(* Logix 5000 project; controller FV vendor 1 type 14 code 217 rev 31.11; software revision 31.00; part 27 of 63 *)
(* tags used below, declared in another part *)
   Alarm_Reset : BOOL;
   Default_Check_Time : DINT;
   Dummy : BOOL;
   FR_B230 : INT[255];   // FLOW_BITS Flow Meter Bits
   FR_B240 : INT[255];   // DEBOUNCE Debounce Flags
   FR_B246 : INT[255];   // V_REVERSE Flags for reversing contol action
   FR_B247 : INT[255];   // CHECKWORD Simulation Flags for Checkwords
   FR_B248 : INT[255];   // FORCE ON Force On Flags
   FR_B249 : INT[255];   // FORCE_OFF NOT Force Off Flags
   FR_B3 : INT[255];   // BINARY
   FR_bit_data_file_address : DINT;
   FR_bit_file_bit_offset : DINT;
   FR_bit_file_word_offset : DINT;
   FR_bit_offset : DINT;
   FR_bit_value_to_set : DINT;
   FR_data_file_address : DINT;
   FR_FRV1_AV01 : PlantItem;   // FRV1_AV01
   FR_FRV1_AV01_ALARM : ALARM_DIGITAL;
   FR_FRV1_AV01_C : ALIAS FOR RIO_Rack_2:4:I.Data.15;
   FR_FRV1_AV01_DR : ALIAS FOR RIO_Rack_2:5:O.Data.7;
   FR_FRV1_AV01_O : ALIAS FOR RIO_Rack_2:4:I.Data.11;
   FR_FV26_AV01 : PlantItem;   // FV26_AV01
   FR_FV26_AV01_ALARM : ALARM_DIGITAL;
   FR_FV26_AV01_C : ALIAS FOR RIO_Rack_2:4:I.Data.20;
   FR_FV26_AV01_O : ALIAS FOR RIO_Rack_2:4:I.Data.16;
   FR_FV26_AV01_RDR : ALIAS FOR RIO_Rack_2:5:O.Data.8;
   FR_FV26_AV04 : PlantItem;   // FV26_AV04
   FR_FV26_AV04_ALARM : ALARM_DIGITAL;
   FR_FV26_AV04_C : ALIAS FOR RIO_Rack_2:4:I.Data.21;
   FR_FV26_AV04_DR : ALIAS FOR RIO_Rack_2:5:O.Data.9;
   FR_FV26_AV04_O : ALIAS FOR RIO_Rack_2:4:I.Data.17;
   FR_FV26_AV05 : PlantItem;   // FV26_AV05
   FR_FV26_AV05_ALARM : ALARM_DIGITAL;
   FR_FV26_AV05_C : ALIAS FOR RIO_Rack_2:4:I.Data.22;
   FR_FV26_AV05_DR : ALIAS FOR RIO_Rack_2:5:O.Data.10;
   FR_FV26_AV05_O : ALIAS FOR RIO_Rack_2:4:I.Data.18;
   FR_FV26_AV06 : PlantItem;   // FV26_AV06
   FR_FV26_AV06_ALARM : ALARM_DIGITAL;
   FR_FV26_AV06_C : ALIAS FOR RIO_Rack_2:4:I.Data.23;
   FR_FV26_AV06_DR : ALIAS FOR RIO_Rack_2:5:O.Data.11;
   FR_FV26_AV06_O : ALIAS FOR RIO_Rack_2:4:I.Data.19;
   FR_FV26_AV07 : PlantItem;   // FV26_AV07
   FR_FV26_AV07_ALARM : ALARM_DIGITAL;
   FR_FV26_AV07_C : ALIAS FOR RIO_Rack_2:4:I.Data.28;
   FR_FV26_AV07_DR : ALIAS FOR RIO_Rack_2:5:O.Data.12;
   FR_FV26_AV07_O : ALIAS FOR RIO_Rack_2:4:I.Data.24;
   FR_FV27_AV01 : PlantItem;   // FV27_AV01
   FR_FV27_AV01_ALARM : ALARM_DIGITAL;
   FR_FV27_AV01_C : ALIAS FOR RIO_Rack_2:4:I.Data.29;
   FR_FV27_AV01_O : ALIAS FOR RIO_Rack_2:4:I.Data.25;
   FR_FV27_AV01_RDR : ALIAS FOR RIO_Rack_2:5:O.Data.13;
   FR_FV27_AV04 : PlantItem;   // FV27_AV04
   FR_FV27_AV04_ALARM : ALARM_DIGITAL;
   FR_FV27_AV04_C : ALIAS FOR RIO_Rack_2:4:I.Data.30;
   FR_FV27_AV04_DR : ALIAS FOR RIO_Rack_2:5:O.Data.14;
   FR_FV27_AV04_O : ALIAS FOR RIO_Rack_2:4:I.Data.26;
   FR_FV27_AV05 : PlantItem;   // FV27_AV05
   FR_FV27_AV05_ALARM : ALARM_DIGITAL;
   FR_FV27_AV05_C : ALIAS FOR RIO_Rack_2:4:I.Data.31;
   FR_FV27_AV05_DR : ALIAS FOR RIO_Rack_2:5:O.Data.15;
   FR_FV27_AV05_O : ALIAS FOR RIO_Rack_2:4:I.Data.27;
   FR_FV27_AV06 : PlantItem;   // FV27_AV06
   FR_FV27_AV06_ALARM : ALARM_DIGITAL;
   FR_FV27_AV06_C : ALIAS FOR RIO_Rack_2:6:I.Data.4;
   FR_FV27_AV06_DR : ALIAS FOR RIO_Rack_2:5:O.Data.16;
   FR_FV27_AV06_O : ALIAS FOR RIO_Rack_2:6:I.Data.0;
   FR_FV27_AV07 : PlantItem;   // FV27_AV07
   FR_FV27_AV07_ALARM : ALARM_DIGITAL;
   FR_FV27_AV07_C : ALIAS FOR RIO_Rack_2:6:I.Data.5;
   FR_FV27_AV07_DR : ALIAS FOR RIO_Rack_2:5:O.Data.17;
   FR_FV27_AV07_O : ALIAS FOR RIO_Rack_2:6:I.Data.1;
   FR_N10 : INT[265];   // FV_AGING Comms to FV Aging PL C
   FR_N100 : INT[265];   // FV FILLING
   FR_N110 : INT[265];   // GREEN BEER Green Beer Main
   FR_N120 : INT[265];   // YEAST CROP Yeast Cropping Main
   FR_N13 : INT[265];   // MV_ROUTE Comms to MV Routing PLC
   FR_N130 : INT[265];   // FILTRATE Filtrate Return
   FR_N14 : INT[265];   // MVFV CIP Comms to MVFV CIP Un it PLC
   FR_N140 : INT[265];   // CIP
   FR_N142 : INT[265];   // CIP
   FR_N143 : INT[265];   // CIP
   FR_N150 : INT[265];   // Original N File From SLC, No Description Available
   FR_N160 : INT[265];   // VESSEL Vessel Working Direc tory
   FR_N170 : INT[265];   // Original N File From SLC, No Description Available
   FR_N180 : INT[265];   // Original N File From SLC, No Description Available
   FR_N198 : INT[265];   // Original N File From SLC, No Description Available
   FR_N20 : INT[265];   // GENERAL General Purpose Setp oints
   FR_N200 : INT[265];   // ANALOG_IN Analog Inputs
   FR_N201 : INT[265];   // Original N File From SLC, No Description Available
   FR_N207 : INT[265];   // Original N File From SLC, No Description Available
   FR_N21 : INT[265];   // CHASE_V FV Filling Beer Chas e Volumes
   FR_N210 : INT[265];   // ANALOG_OUT Analog Outputs
   FR_N220 : INT[265];   // CHECKLIST Checklist Loop Contr ollers
   FR_N225 : INT[265];   // Original N File From SLC, No Description Available
   FR_N226 : INT[265];   // Original N File From SLC, No Description Available
   FR_N245 : INT[265];   // CHECKWORD Checkword Loop Contr ol
   FR_N252 : INT[265];   // OUTPUT_PTR Checkword Pointers t o output flags in B2 50
   FR_N253 : INT[265];   // EN_POINT Pointers to energise d input flags in B25 1
   FR_N254 : INT[265];   // DEN_POINT Pointers to deenergi sed input flags in B 251
   FR_N255 : INT[265];   // CHECKWORDS
   FR_N26 : INT[265];   // FV26
   FR_N27 : INT[265];   // FV27
   FR_N28 : INT[265];   // FV28
   FR_N29 : INT[265];   // FV29
   FR_N30 : INT[265];   // FV30
   FR_N31 : INT[265];   // FV31
   FR_N36 : INT[265];   // Original N File From SLC, No Description Available
   FR_N37 : INT[265];   // Original N File From SLC, No Description Available
   FR_N46 : INT[265];   // Original N File From SLC, No Description Available
   FR_N47 : INT[265];   // Original N File From SLC, No Description Available
   FR_N7 : INT[265];   // INTEGER
   FR_N99 : INT[265];   // COMMENT Comment Lines
   FR_value_to_set : DINT;
   FR_VB1_AV01 : PlantItem;   // VB1_AV01
   FR_VB1_AV01_ALARM : ALARM_DIGITAL;
   FR_VB1_AV01_C : ALIAS FOR RIO_Rack_2:6:I.Data.6;
   FR_VB1_AV01_DR : ALIAS FOR RIO_Rack_2:5:O.Data.18;
   FR_VB1_AV01_O : ALIAS FOR RIO_Rack_2:6:I.Data.2;
   FR_VB1_AV02 : PlantItem;   // VB1_AV02
   FR_VB1_AV02_ALARM : ALARM_DIGITAL;
   FR_VB1_AV02_C : ALIAS FOR RIO_Rack_2:6:I.Data.7;
   FR_VB1_AV02_DR : ALIAS FOR RIO_Rack_2:5:O.Data.19;
   FR_VB1_AV02_O : ALIAS FOR RIO_Rack_2:6:I.Data.3;
   FR_VB1_AV03 : PlantItem;   // VB1_AV03
   FR_VB1_AV03_ALARM : ALARM_DIGITAL;
   FR_VB1_AV03_C : ALIAS FOR RIO_Rack_2:6:I.Data.12;
   FR_VB1_AV03_DR : ALIAS FOR RIO_Rack_2:5:O.Data.20;
   FR_VB1_AV03_O : ALIAS FOR RIO_Rack_2:6:I.Data.8;
   FR_word_offset : DINT;
   Item_Faults_Are_Latched : BOOL;
   Item_Simulation_Flag : BOOL;
   One_Second_One_Scan : ALIAS FOR One_Second_1_scan;
(* FR_Common, continued *)

ROUTINE FR_Set_NFile_Value   (* ladder *)
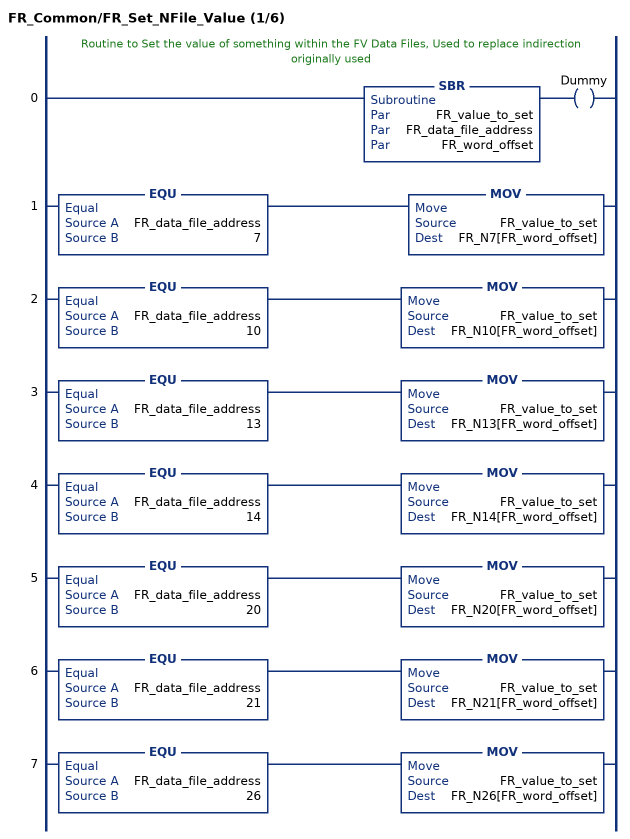
   // Routine to Set the value of something within the FV Data Files, Used to replace indirection originally used
   0: SBR(FR_value_to_set,FR_data_file_address,FR_word_offset)OTE(Dummy);
   1: EQU(FR_data_file_address,7)MOV(FR_value_to_set,FR_N7[FR_word_offset]);
   2: EQU(FR_data_file_address,10)MOV(FR_value_to_set,FR_N10[FR_word_offset]);
   3: EQU(FR_data_file_address,13)MOV(FR_value_to_set,FR_N13[FR_word_offset]);
   4: EQU(FR_data_file_address,14)MOV(FR_value_to_set,FR_N14[FR_word_offset]);
   5: EQU(FR_data_file_address,20)MOV(FR_value_to_set,FR_N20[FR_word_offset]);
   6: EQU(FR_data_file_address,21)MOV(FR_value_to_set,FR_N21[FR_word_offset]);
   7: EQU(FR_data_file_address,26)MOV(FR_value_to_set,FR_N26[FR_word_offset]);
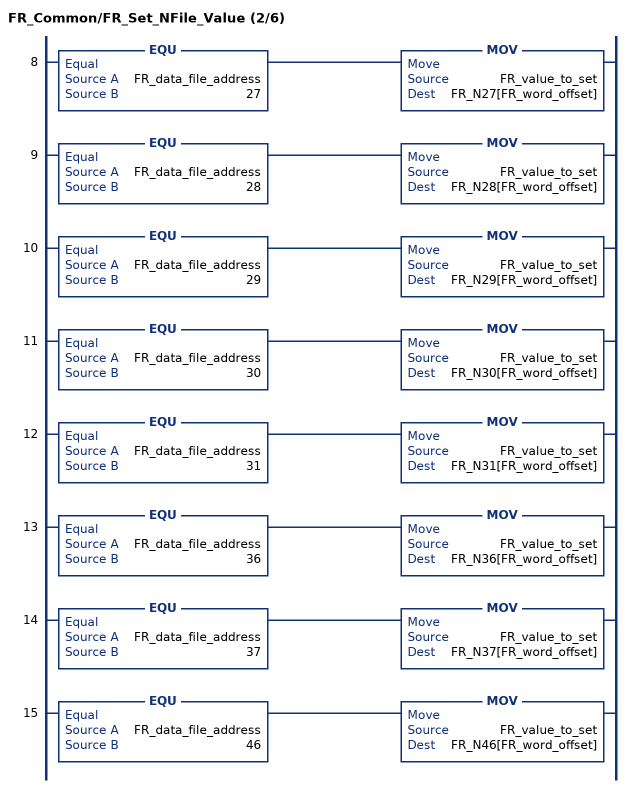
   8: EQU(FR_data_file_address,27)MOV(FR_value_to_set,FR_N27[FR_word_offset]);
   9: EQU(FR_data_file_address,28)MOV(FR_value_to_set,FR_N28[FR_word_offset]);
   10: EQU(FR_data_file_address,29)MOV(FR_value_to_set,FR_N29[FR_word_offset]);
   11: EQU(FR_data_file_address,30)MOV(FR_value_to_set,FR_N30[FR_word_offset]);
   12: EQU(FR_data_file_address,31)MOV(FR_value_to_set,FR_N31[FR_word_offset]);
   13: EQU(FR_data_file_address,36)MOV(FR_value_to_set,FR_N36[FR_word_offset]);
   14: EQU(FR_data_file_address,37)MOV(FR_value_to_set,FR_N37[FR_word_offset]);
   15: EQU(FR_data_file_address,46)MOV(FR_value_to_set,FR_N46[FR_word_offset]);
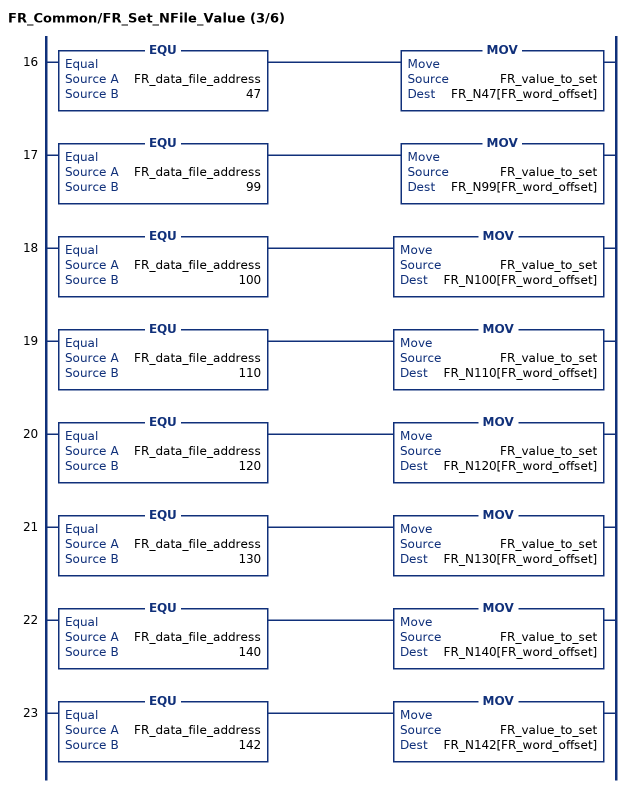
   16: EQU(FR_data_file_address,47)MOV(FR_value_to_set,FR_N47[FR_word_offset]);
   17: EQU(FR_data_file_address,99)MOV(FR_value_to_set,FR_N99[FR_word_offset]);
   18: EQU(FR_data_file_address,100)MOV(FR_value_to_set,FR_N100[FR_word_offset]);
   19: EQU(FR_data_file_address,110)MOV(FR_value_to_set,FR_N110[FR_word_offset]);
   20: EQU(FR_data_file_address,120)MOV(FR_value_to_set,FR_N120[FR_word_offset]);
   21: EQU(FR_data_file_address,130)MOV(FR_value_to_set,FR_N130[FR_word_offset]);
   22: EQU(FR_data_file_address,140)MOV(FR_value_to_set,FR_N140[FR_word_offset]);
   23: EQU(FR_data_file_address,142)MOV(FR_value_to_set,FR_N142[FR_word_offset]);
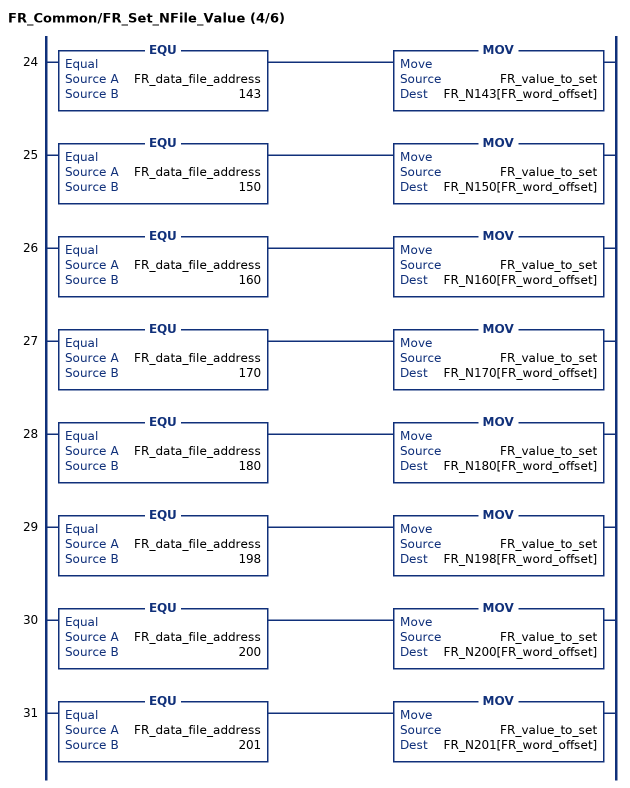
   24: EQU(FR_data_file_address,143)MOV(FR_value_to_set,FR_N143[FR_word_offset]);
   25: EQU(FR_data_file_address,150)MOV(FR_value_to_set,FR_N150[FR_word_offset]);
   26: EQU(FR_data_file_address,160)MOV(FR_value_to_set,FR_N160[FR_word_offset]);
   27: EQU(FR_data_file_address,170)MOV(FR_value_to_set,FR_N170[FR_word_offset]);
   28: EQU(FR_data_file_address,180)MOV(FR_value_to_set,FR_N180[FR_word_offset]);
   29: EQU(FR_data_file_address,198)MOV(FR_value_to_set,FR_N198[FR_word_offset]);
   30: EQU(FR_data_file_address,200)MOV(FR_value_to_set,FR_N200[FR_word_offset]);
   31: EQU(FR_data_file_address,201)MOV(FR_value_to_set,FR_N201[FR_word_offset]);
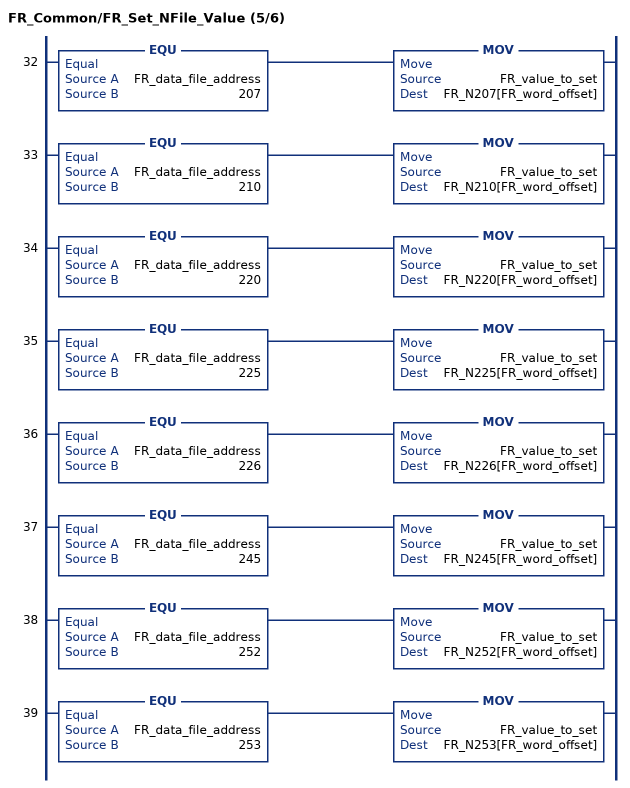
   32: EQU(FR_data_file_address,207)MOV(FR_value_to_set,FR_N207[FR_word_offset]);
   33: EQU(FR_data_file_address,210)MOV(FR_value_to_set,FR_N210[FR_word_offset]);
   34: EQU(FR_data_file_address,220)MOV(FR_value_to_set,FR_N220[FR_word_offset]);
   35: EQU(FR_data_file_address,225)MOV(FR_value_to_set,FR_N225[FR_word_offset]);
   36: EQU(FR_data_file_address,226)MOV(FR_value_to_set,FR_N226[FR_word_offset]);
   37: EQU(FR_data_file_address,245)MOV(FR_value_to_set,FR_N245[FR_word_offset]);
   38: EQU(FR_data_file_address,252)MOV(FR_value_to_set,FR_N252[FR_word_offset]);
   39: EQU(FR_data_file_address,253)MOV(FR_value_to_set,FR_N253[FR_word_offset]);
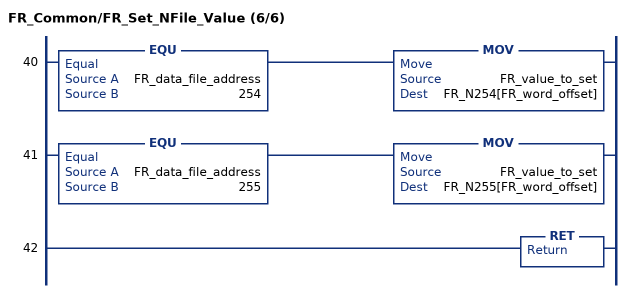
   40: EQU(FR_data_file_address,254)MOV(FR_value_to_set,FR_N254[FR_word_offset]);
   41: EQU(FR_data_file_address,255)MOV(FR_value_to_set,FR_N255[FR_word_offset]);
   42: RET();
END_ROUTINE

ROUTINE FR_SetBitFile_Value   (* ladder *)
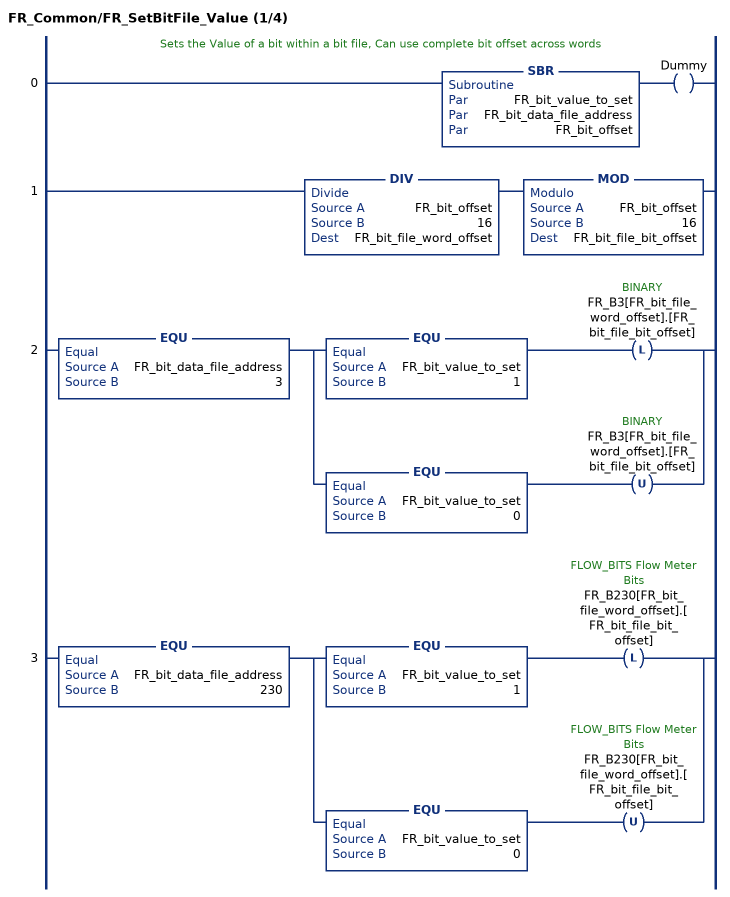
   // Sets the Value of a bit within a bit file, Can use complete bit offset across words
   0: SBR(FR_bit_value_to_set,FR_bit_data_file_address,FR_bit_offset)OTE(Dummy);
   1: DIV(FR_bit_offset,16,FR_bit_file_word_offset)MOD(FR_bit_offset,16,FR_bit_file_bit_offset);
   2: EQU(FR_bit_data_file_address,3)[EQU(FR_bit_value_to_set,1) OTL(FR_B3[FR_bit_file_word_offset].[FR_bit_file_bit_offset]) ,EQU(FR_bit_value_to_set,0) OTU(FR_B3[FR_bit_file_word_offset].[FR_bit_file_bit_offset]) ];
   3: EQU(FR_bit_data_file_address,230)[EQU(FR_bit_value_to_set,1) OTL(FR_B230[FR_bit_file_word_offset].[FR_bit_file_bit_offset]) ,EQU(FR_bit_value_to_set,0) OTU(FR_B230[FR_bit_file_word_offset].[FR_bit_file_bit_offset]) ];
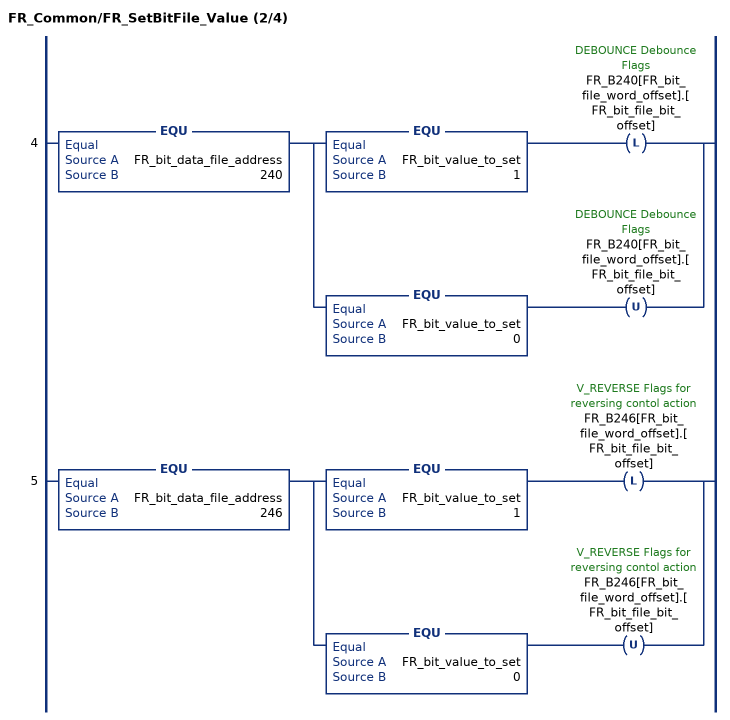
   4: EQU(FR_bit_data_file_address,240)[EQU(FR_bit_value_to_set,1) OTL(FR_B240[FR_bit_file_word_offset].[FR_bit_file_bit_offset]) ,EQU(FR_bit_value_to_set,0) OTU(FR_B240[FR_bit_file_word_offset].[FR_bit_file_bit_offset]) ];
   5: EQU(FR_bit_data_file_address,246)[EQU(FR_bit_value_to_set,1) OTL(FR_B246[FR_bit_file_word_offset].[FR_bit_file_bit_offset]) ,EQU(FR_bit_value_to_set,0) OTU(FR_B246[FR_bit_file_word_offset].[FR_bit_file_bit_offset]) ];
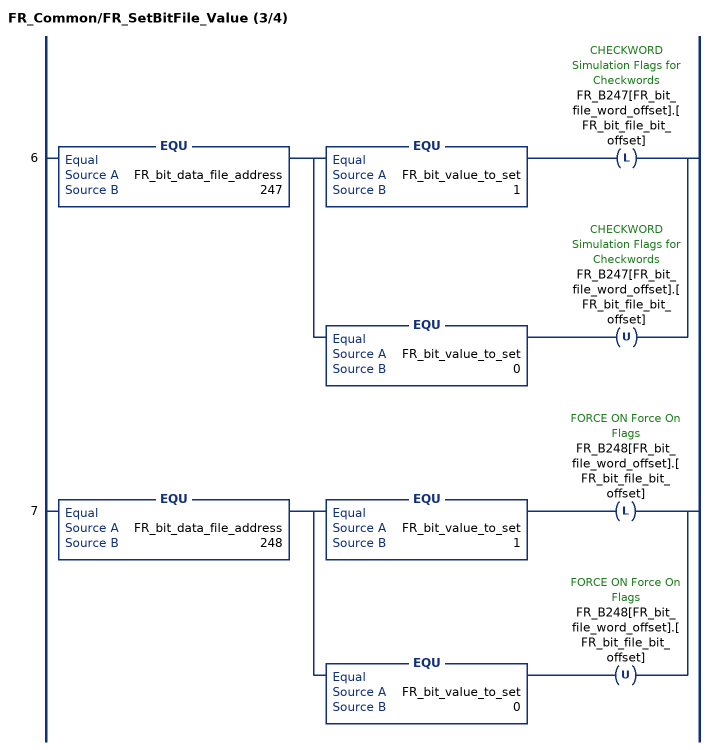
   6: EQU(FR_bit_data_file_address,247)[EQU(FR_bit_value_to_set,1) OTL(FR_B247[FR_bit_file_word_offset].[FR_bit_file_bit_offset]) ,EQU(FR_bit_value_to_set,0) OTU(FR_B247[FR_bit_file_word_offset].[FR_bit_file_bit_offset]) ];
   7: EQU(FR_bit_data_file_address,248)[EQU(FR_bit_value_to_set,1) OTL(FR_B248[FR_bit_file_word_offset].[FR_bit_file_bit_offset]) ,EQU(FR_bit_value_to_set,0) OTU(FR_B248[FR_bit_file_word_offset].[FR_bit_file_bit_offset]) ];
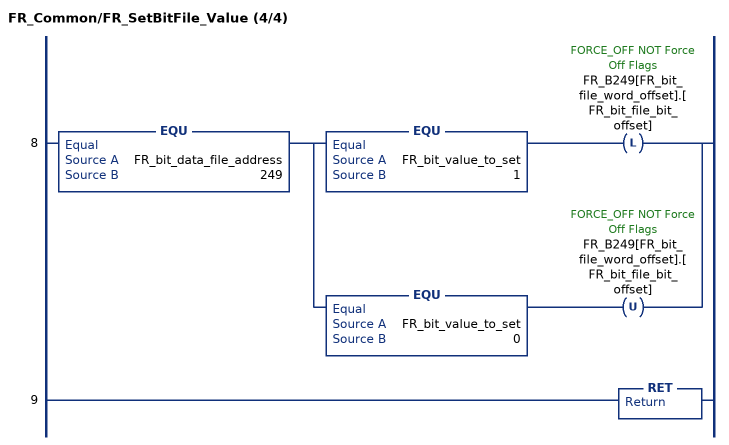
   8: EQU(FR_bit_data_file_address,249)[EQU(FR_bit_value_to_set,1) OTL(FR_B249[FR_bit_file_word_offset].[FR_bit_file_bit_offset]) ,EQU(FR_bit_value_to_set,0) OTU(FR_B249[FR_bit_file_word_offset].[FR_bit_file_bit_offset]) ];
   9: RET();
END_ROUTINE

ROUTINE FR_Valves   (* ladder *)
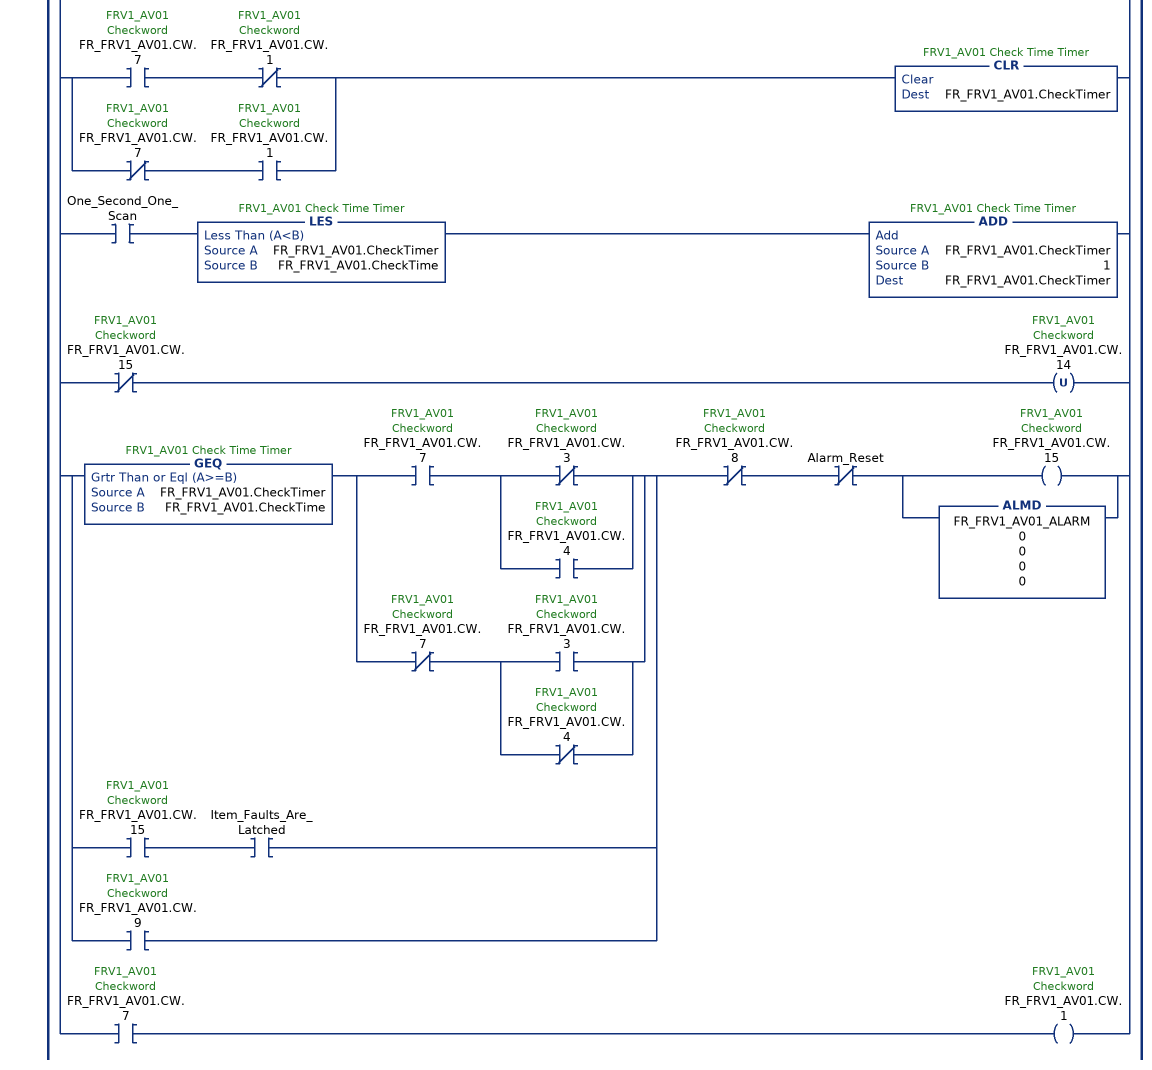
   0: [NEQ(FR_FRV1_AV01.DriveBits,0) OTE(FR_FRV1_AV01.CW.0) ,[XIC(FR_FRV1_AV01.CW.0) XIO(FR_FRV1_AV01.CW.6) ,XIC(FR_FRV1_AV01.CW.5) XIC(FR_FRV1_AV01.CW.6) ] OTE(FR_FRV1_AV01.CW.7) ,XIC(FR_FRV1_AV01.CW.7) OTE(FR_FRV1_AV01_DR) ,XIC(S:FS) [OTU(FR_FRV1_AV01.CW.6) ,LEQ(FR_FRV1_AV01.CheckTime,0) MOV(Default_Check_Time,FR_FRV1_AV01.CheckTime) ] ,[[XIC(FR_FRV1_AV01_O) XIO(Item_Simulation_Flag) ,XIC(Item_Simulation_Flag) XIC(FR_FRV1_AV01.CW.7) XIO(FR_FRV1_AV01.CW.2) ] OTE(FR_FRV1_AV01.CW.3) ,[XIC(FR_FRV1_AV01_C) XIO(Item_Simulation_Flag) ,XIC(Item_Simulation_Flag) XIO(FR_FRV1_AV01.CW.7) XIO(FR_FRV1_AV01.CW.2) ] OTE(FR_FRV1_AV01.CW.4) ] ,[XIC(FR_FRV1_AV01.CW.7) XIO(FR_FRV1_AV01.CW.1) ,XIO(FR_FRV1_AV01.CW.7) XIC(FR_FRV1_AV01.CW.1) ] CLR(FR_FRV1_AV01.CheckTimer) ,XIC(One_Second_One_Scan) LES(FR_FRV1_AV01.CheckTimer,FR_FRV1_AV01.CheckTime) ADD(FR_FRV1_AV01.CheckTimer,1,FR_FRV1_AV01.CheckTimer) ,XIO(FR_FRV1_AV01.CW.15) OTU(FR_FRV1_AV01.CW.14) ,[GEQ(FR_FRV1_AV01.CheckTimer,FR_FRV1_AV01.CheckTime) [XIC(FR_FRV1_AV01.CW.7) [XIO(FR_FRV1_AV01.CW.3) ,XIC(FR_FRV1_AV01.CW.4) ] ,XIO(FR_FRV1_AV01.CW.7) [XIC(FR_FRV1_AV01.CW.3) ,XIO(FR_FRV1_AV01.CW.4) ] ] ,XIC(FR_FRV1_AV01.CW.15) XIC(Item_Faults_Are_Latched) ,XIC(FR_FRV1_AV01.CW.9) ] XIO(FR_FRV1_AV01.CW.8) XIO(Alarm_Reset) [OTE(FR_FRV1_AV01.CW.15) ,ALMD(FR_FRV1_AV01_ALARM,0,0,0,0) ] ,XIC(FR_FRV1_AV01.CW.7) OTE(FR_FRV1_AV01.CW.1) ];
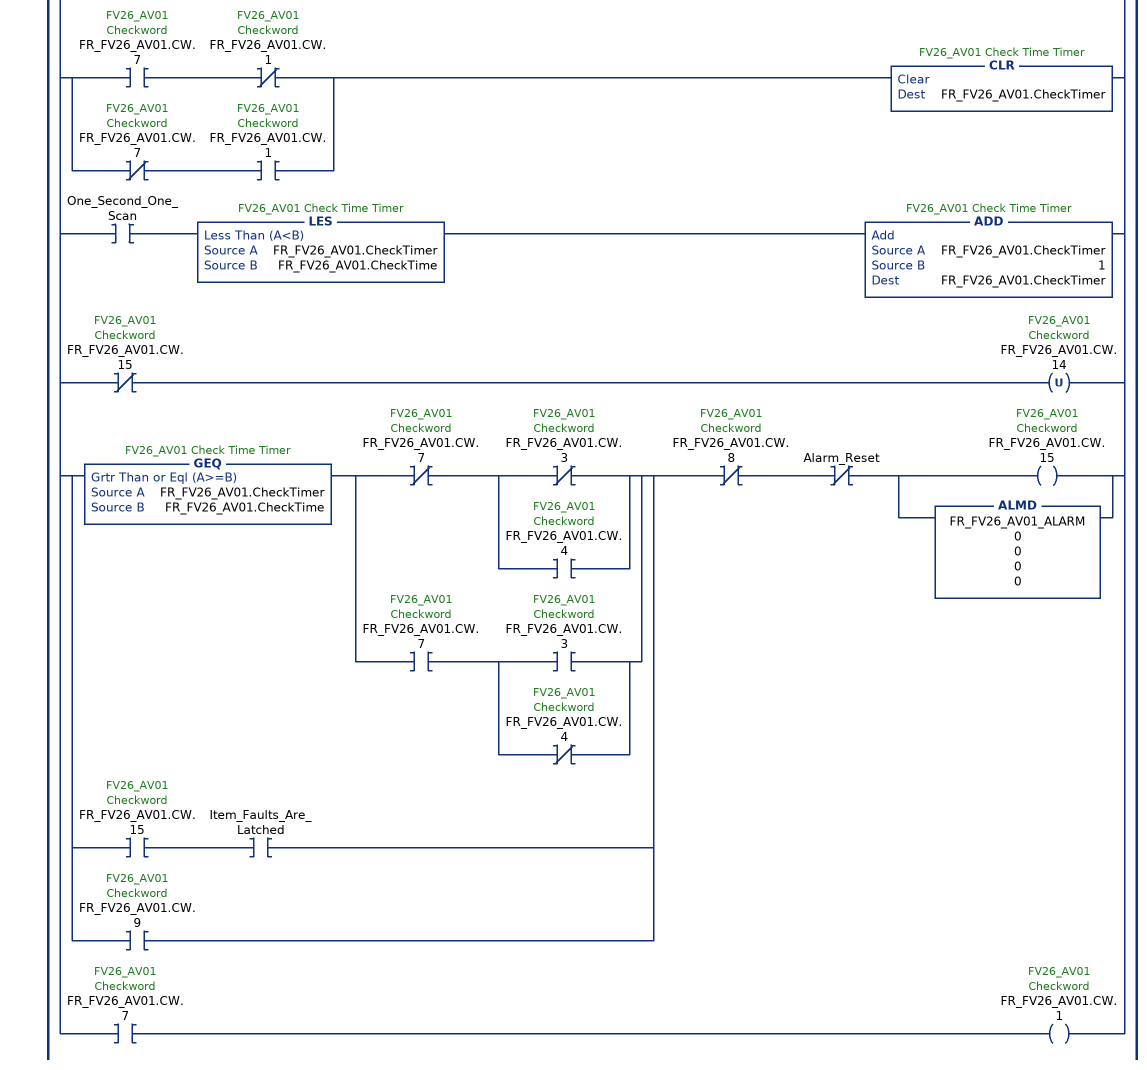
   1: [NEQ(FR_FV26_AV01.DriveBits,0) OTE(FR_FV26_AV01.CW.0) ,[XIC(FR_FV26_AV01.CW.0) XIO(FR_FV26_AV01.CW.6) ,XIC(FR_FV26_AV01.CW.5) XIC(FR_FV26_AV01.CW.6) ] OTE(FR_FV26_AV01.CW.7) ,XIC(FR_FV26_AV01.CW.7) OTE(FR_FV26_AV01_RDR) ,XIC(S:FS) [OTU(FR_FV26_AV01.CW.6) ,LEQ(FR_FV26_AV01.CheckTime,0) MOV(Default_Check_Time,FR_FV26_AV01.CheckTime) ] ,[[XIC(FR_FV26_AV01_C) XIO(Item_Simulation_Flag) ,XIC(Item_Simulation_Flag) XIO(FR_FV26_AV01.CW.7) XIO(FR_FV26_AV01.CW.2) ] OTE(FR_FV26_AV01.CW.3) ,[XIC(FR_FV26_AV01_O) XIO(Item_Simulation_Flag) ,XIC(Item_Simulation_Flag) XIC(FR_FV26_AV01.CW.7) XIO(FR_FV26_AV01.CW.2) ] OTE(FR_FV26_AV01.CW.4) ] ,[XIC(FR_FV26_AV01.CW.7) XIO(FR_FV26_AV01.CW.1) ,XIO(FR_FV26_AV01.CW.7) XIC(FR_FV26_AV01.CW.1) ] CLR(FR_FV26_AV01.CheckTimer) ,XIC(One_Second_One_Scan) LES(FR_FV26_AV01.CheckTimer,FR_FV26_AV01.CheckTime) ADD(FR_FV26_AV01.CheckTimer,1,FR_FV26_AV01.CheckTimer) ,XIO(FR_FV26_AV01.CW.15) OTU(FR_FV26_AV01.CW.14) ,[GEQ(FR_FV26_AV01.CheckTimer,FR_FV26_AV01.CheckTime) [XIO(FR_FV26_AV01.CW.7) [XIO(FR_FV26_AV01.CW.3) ,XIC(FR_FV26_AV01.CW.4) ] ,XIC(FR_FV26_AV01.CW.7) [XIC(FR_FV26_AV01.CW.3) ,XIO(FR_FV26_AV01.CW.4) ] ] ,XIC(FR_FV26_AV01.CW.15) XIC(Item_Faults_Are_Latched) ,XIC(FR_FV26_AV01.CW.9) ] XIO(FR_FV26_AV01.CW.8) XIO(Alarm_Reset) [OTE(FR_FV26_AV01.CW.15) ,ALMD(FR_FV26_AV01_ALARM,0,0,0,0) ] ,XIC(FR_FV26_AV01.CW.7) OTE(FR_FV26_AV01.CW.1) ];
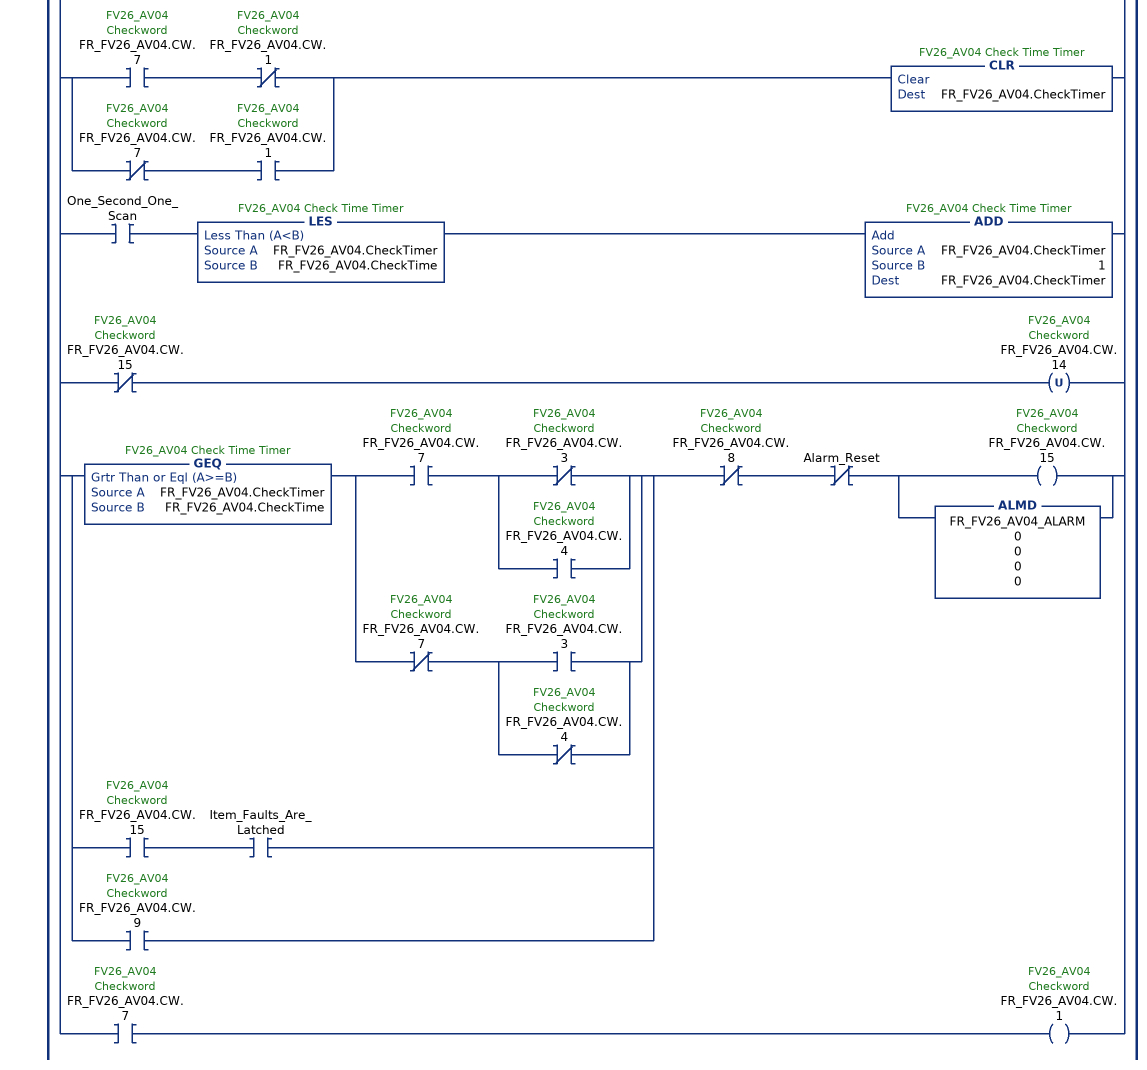
   2: [NEQ(FR_FV26_AV04.DriveBits,0) OTE(FR_FV26_AV04.CW.0) ,[XIC(FR_FV26_AV04.CW.0) XIO(FR_FV26_AV04.CW.6) ,XIC(FR_FV26_AV04.CW.5) XIC(FR_FV26_AV04.CW.6) ] OTE(FR_FV26_AV04.CW.7) ,XIC(FR_FV26_AV04.CW.7) OTE(FR_FV26_AV04_DR) ,XIC(S:FS) [OTU(FR_FV26_AV04.CW.6) ,LEQ(FR_FV26_AV04.CheckTime,0) MOV(Default_Check_Time,FR_FV26_AV04.CheckTime) ] ,[[XIC(FR_FV26_AV04_O) XIO(Item_Simulation_Flag) ,XIC(Item_Simulation_Flag) XIC(FR_FV26_AV04.CW.7) XIO(FR_FV26_AV04.CW.2) ] OTE(FR_FV26_AV04.CW.3) ,[XIC(FR_FV26_AV04_C) XIO(Item_Simulation_Flag) ,XIC(Item_Simulation_Flag) XIO(FR_FV26_AV04.CW.7) XIO(FR_FV26_AV04.CW.2) ] OTE(FR_FV26_AV04.CW.4) ] ,[XIC(FR_FV26_AV04.CW.7) XIO(FR_FV26_AV04.CW.1) ,XIO(FR_FV26_AV04.CW.7) XIC(FR_FV26_AV04.CW.1) ] CLR(FR_FV26_AV04.CheckTimer) ,XIC(One_Second_One_Scan) LES(FR_FV26_AV04.CheckTimer,FR_FV26_AV04.CheckTime) ADD(FR_FV26_AV04.CheckTimer,1,FR_FV26_AV04.CheckTimer) ,XIO(FR_FV26_AV04.CW.15) OTU(FR_FV26_AV04.CW.14) ,[GEQ(FR_FV26_AV04.CheckTimer,FR_FV26_AV04.CheckTime) [XIC(FR_FV26_AV04.CW.7) [XIO(FR_FV26_AV04.CW.3) ,XIC(FR_FV26_AV04.CW.4) ] ,XIO(FR_FV26_AV04.CW.7) [XIC(FR_FV26_AV04.CW.3) ,XIO(FR_FV26_AV04.CW.4) ] ] ,XIC(FR_FV26_AV04.CW.15) XIC(Item_Faults_Are_Latched) ,XIC(FR_FV26_AV04.CW.9) ] XIO(FR_FV26_AV04.CW.8) XIO(Alarm_Reset) [OTE(FR_FV26_AV04.CW.15) ,ALMD(FR_FV26_AV04_ALARM,0,0,0,0) ] ,XIC(FR_FV26_AV04.CW.7) OTE(FR_FV26_AV04.CW.1) ];
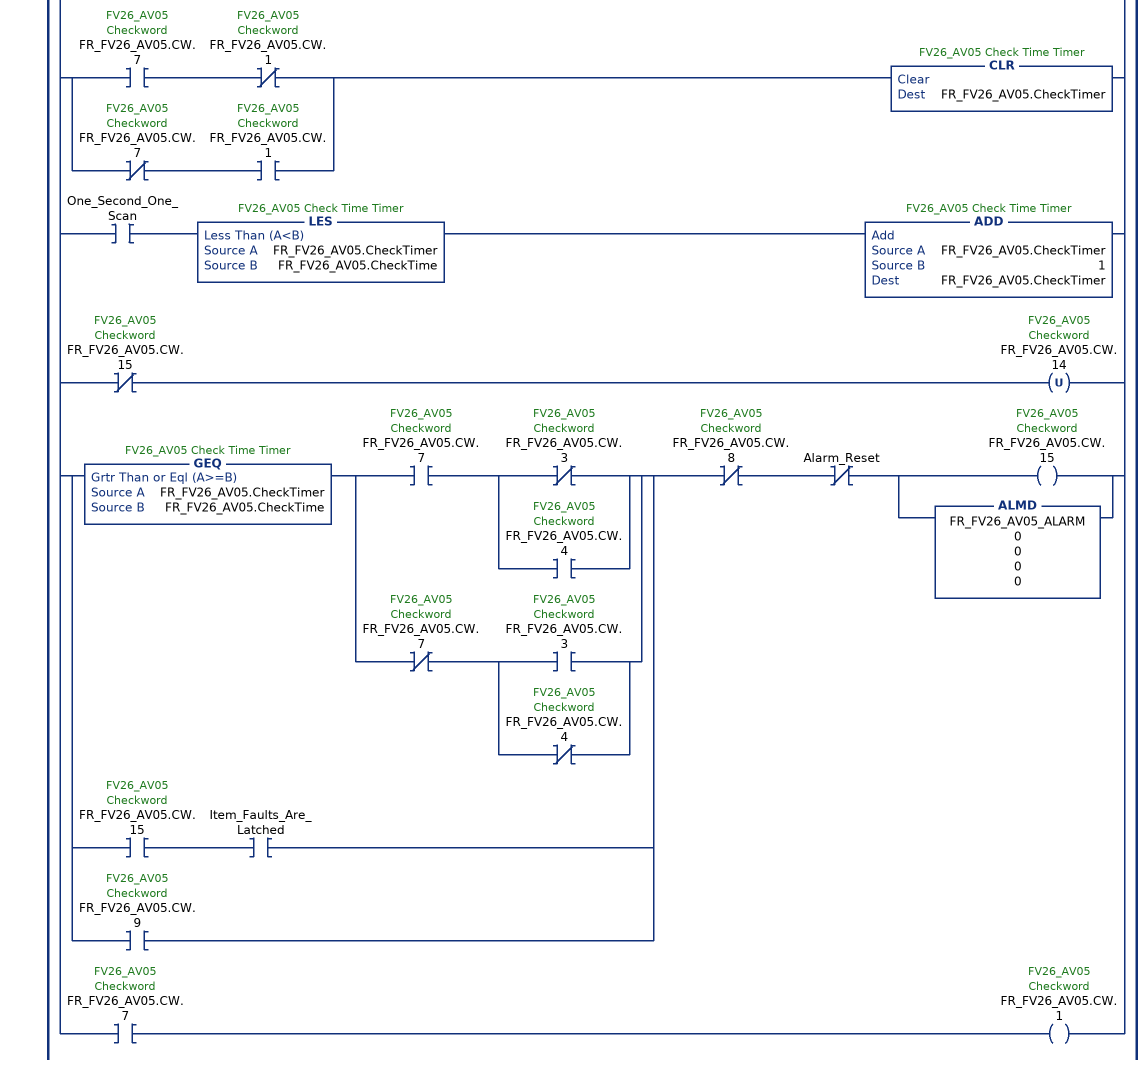
   3: [NEQ(FR_FV26_AV05.DriveBits,0) OTE(FR_FV26_AV05.CW.0) ,[XIC(FR_FV26_AV05.CW.0) XIO(FR_FV26_AV05.CW.6) ,XIC(FR_FV26_AV05.CW.5) XIC(FR_FV26_AV05.CW.6) ] OTE(FR_FV26_AV05.CW.7) ,XIC(FR_FV26_AV05.CW.7) OTE(FR_FV26_AV05_DR) ,XIC(S:FS) [OTU(FR_FV26_AV05.CW.6) ,LEQ(FR_FV26_AV05.CheckTime,0) MOV(Default_Check_Time,FR_FV26_AV05.CheckTime) ] ,[[XIC(FR_FV26_AV05_O) XIO(Item_Simulation_Flag) ,XIC(Item_Simulation_Flag) XIC(FR_FV26_AV05.CW.7) XIO(FR_FV26_AV05.CW.2) ] OTE(FR_FV26_AV05.CW.3) ,[XIC(FR_FV26_AV05_C) XIO(Item_Simulation_Flag) ,XIC(Item_Simulation_Flag) XIO(FR_FV26_AV05.CW.7) XIO(FR_FV26_AV05.CW.2) ] OTE(FR_FV26_AV05.CW.4) ] ,[XIC(FR_FV26_AV05.CW.7) XIO(FR_FV26_AV05.CW.1) ,XIO(FR_FV26_AV05.CW.7) XIC(FR_FV26_AV05.CW.1) ] CLR(FR_FV26_AV05.CheckTimer) ,XIC(One_Second_One_Scan) LES(FR_FV26_AV05.CheckTimer,FR_FV26_AV05.CheckTime) ADD(FR_FV26_AV05.CheckTimer,1,FR_FV26_AV05.CheckTimer) ,XIO(FR_FV26_AV05.CW.15) OTU(FR_FV26_AV05.CW.14) ,[GEQ(FR_FV26_AV05.CheckTimer,FR_FV26_AV05.CheckTime) [XIC(FR_FV26_AV05.CW.7) [XIO(FR_FV26_AV05.CW.3) ,XIC(FR_FV26_AV05.CW.4) ] ,XIO(FR_FV26_AV05.CW.7) [XIC(FR_FV26_AV05.CW.3) ,XIO(FR_FV26_AV05.CW.4) ] ] ,XIC(FR_FV26_AV05.CW.15) XIC(Item_Faults_Are_Latched) ,XIC(FR_FV26_AV05.CW.9) ] XIO(FR_FV26_AV05.CW.8) XIO(Alarm_Reset) [OTE(FR_FV26_AV05.CW.15) ,ALMD(FR_FV26_AV05_ALARM,0,0,0,0) ] ,XIC(FR_FV26_AV05.CW.7) OTE(FR_FV26_AV05.CW.1) ];